// TIA Portal project "Mixing_Process" (V19)
// Mixing of two ingredients process

(* hardware
DEVICE "S7-1200 station_1"  S7-1200 Station
   slot 0: "Rack_0"  S7-1200 Rack  Rack  V1.0
   slot 1: "PLC_1"  CPU 1212C AC/DC/Rly  6ES7 212-1BE40-0XB0  V4.6
DEVICE "HMI_1"  TP1200 Comfort
   slot 0: "HMI_1"  TP1200 Comfort  6AV2 124-0MC01-0AX0  17.0.0.0
   slot 1: "HMI_RT_1"  TP1200 Comfort  6AV2 124-0MC01-0AX0  17.0.0.0
   slot 5: "HMI_1.IE_CP_1"  PROFINET Interface  17.0.0.0
      slot 1: "PROFINET Interface_1"  PROFINET Interface
         slot 1: "Port_1"  Port
         slot 2: "Port_2"  Port
   slot 7: "HMI_1.MPI/DP_CP_1"  MPI/DP Interface  17.0.0.0
*)

// ===== PLC "PLC_1"  CPU 1212C AC/DC/Rly =====

VAR_GLOBAL   // PLC tag table "Inputs"
   "E_Stop" AT %I0.0 : Bool;   // Stop mushroom
   "Pb_Stop" AT %I0.1 : Bool;   // Pushbutton Stop
   "Pb_Start" AT %I0.2 : Bool;   // Pushbutton Start
   "Tank_Empty_Level" AT %I0.3 : Bool;   // Empty level sensor, NO logic
   "Level_A" AT %I0.4 : Bool;   // Level for liquid A, NO logic
   "Level_B" AT %I0.5 : Bool;   // Level for liquid B, NO logic
   "Thermal_Fault" AT %I0.6 : Bool;   // Thermal fault from thermal relay
   "Temp_Alm" AT %I0.7 : Bool;   // Temperature alarm from control temperature
   "Tag_1" AT %M0.0 : Bool;
END_VAR

VAR_GLOBAL   // PLC tag table "Outputs"
   "Motor_Mixer" AT %Q0.0 : Bool;   // Motor mixer
   "Valve_A" AT %Q0.1 : Bool;   // Valve liquid A
   "Valve_B" AT %Q0.2 : Bool;   // Valve liquid B
   "Temp_Relay" AT %Q0.4 : Bool;   // Control relay for temperature signal
   "Valve_C" AT %Q0.5 : Bool;   // Discharge Valve
END_VAR

// folder: DB

DATA_BLOCK "DATA"   // DB1
TITLE = Data blocks for functions
{ S7_Optimized_Access := 'TRUE' }
AUTHOR : Stiven Perez Mora
VERSION : 0.1
   VAR
      Start_Stop : Bool;
      Q_TimeDischarge : Bool;
      E_Discharge : Int;
      Active_Valve_C : Bool;
      E_Active_Valve_C : Bool;
      E_Stop : Bool;
      Pb_Start : Bool;
   END_VAR
BEGIN
END_DATA_BLOCK

DATA_BLOCK "HMI_Data"   // DB4
{ S7_Optimized_Access := 'TRUE' }
VERSION : 0.1
   VAR
      Start_HMI : Bool;
      Stop_HMI : Bool;
      Valve_A : Bool;
      Level_A : Bool;
      Valve_B : Bool;
      Level_B : Bool;
      Valve_C : Bool;
      Motor_Mixer : Bool;
      Temp_Relay : Bool;
      PT_Mixing : Time;   // Miliseconds timer mix
      PT_M_Mxing : Time;   // Minutes timer mix
      ET_Mixing : Time;   // Miliseconds elapsed time
      ET_Mixing_S : Time;   // Seconds elapsed time
      Empty_Level : Bool;
      Empty_Field_Time : Bool;   // Ambar text alert, input mix time
   END_VAR
BEGIN
END_DATA_BLOCK

// folder: System blocks/Program resources

DATA_BLOCK "TimeToWamUp"   // DB2
{ S7_Optimized_Access := 'TRUE' }
AUTHOR : Simatic
FAMILY : IEC
NAME : IEC_TMR
VERSION : 1.0
// stored: InstanceOfName IEC_TIMER
"IEC_TIMER"
BEGIN
END_DATA_BLOCK

DATA_BLOCK "TimeToMixing"   // DB3
{ S7_Optimized_Access := 'TRUE' }
AUTHOR : Simatic
FAMILY : IEC
NAME : IEC_TMR
VERSION : 1.0
// stored: InstanceOfName IEC_TIMER
"IEC_TIMER"
BEGIN
END_DATA_BLOCK

DATA_BLOCK "MixingTime"   // DB5
{ S7_Optimized_Access := 'TRUE' }
AUTHOR : Simatic
FAMILY : IEC
NAME : IEC_TMR
VERSION : 1.0
// stored: InstanceOfName IEC_TIMER
"IEC_TIMER"
BEGIN
END_DATA_BLOCK

// folder: (top level)

ORGANIZATION_BLOCK "Main"   // OB1, LAD, ProgramCycle
TITLE = "Main Program Sweep (Cycle)"
{ S7_Optimized_Access := 'TRUE' }
VERSION : 0.1
   VAR_INPUT
      Initial_Call : Bool;   // Initial call of this OB
      Remanence : Bool;   // =True, if remanent data are available
   END_VAR
BEGIN

REGION Network 1: Block Start or Stop all process
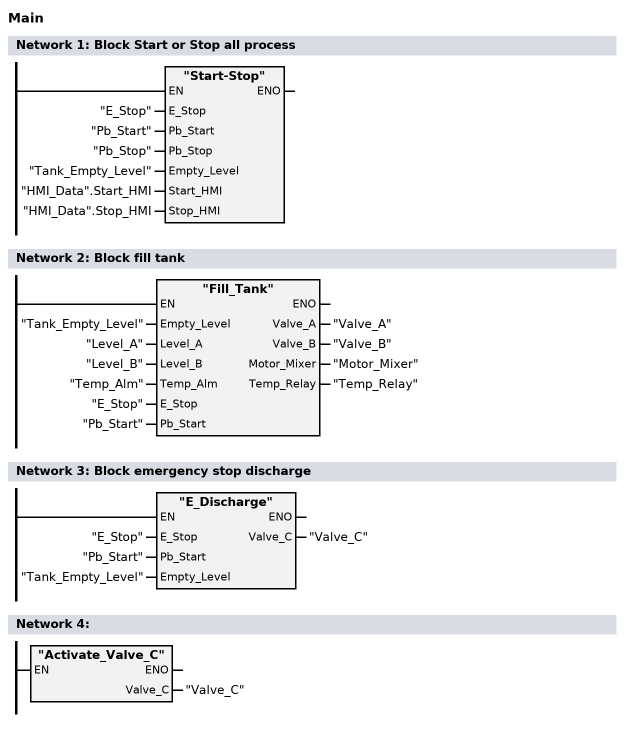
   RUNG wire#powerrail
      "Start-Stop"(E_Stop := "E_Stop", Pb_Start := "Pb_Start", Pb_Stop := "Pb_Stop", Empty_Level := "Tank_Empty_Level", Start_HMI := "HMI_Data".Start_HMI, Stop_HMI := "HMI_Data".Stop_HMI)
   END_RUNG
   // the same network as SCL:
   "Start-Stop"(E_Stop := "E_Stop",
                Pb_Start := "Pb_Start",
                Pb_Stop := "Pb_Stop",
                Empty_Level := "Tank_Empty_Level",
                Start_HMI := "HMI_Data".Start_HMI,
                Stop_HMI := "HMI_Data".Stop_HMI);
END_REGION

REGION Network 2: Block fill tank
   RUNG wire#powerrail
      "Fill_Tank"(Empty_Level := "Tank_Empty_Level", Level_A := "Level_A", Level_B := "Level_B", Temp_Alm := "Temp_Alm", E_Stop := "E_Stop", Pb_Start := "Pb_Start", Valve_A => "Valve_A", Valve_B => "Valve_B", Motor_Mixer => "Motor_Mixer", Temp_Relay => "Temp_Relay")
   END_RUNG
   // the same network as SCL:
   "Fill_Tank"(Empty_Level := "Tank_Empty_Level",
               Level_A := "Level_A",
               Level_B := "Level_B",
               Temp_Alm := "Temp_Alm",
               E_Stop := "E_Stop",
               Pb_Start := "Pb_Start",
               Valve_A => "Valve_A",
               Valve_B => "Valve_B",
               Motor_Mixer => "Motor_Mixer",
               Temp_Relay => "Temp_Relay");
END_REGION

REGION Network 3: Block emergency stop discharge
   RUNG wire#powerrail
      "E_Discharge"(E_Stop := "E_Stop", Pb_Start := "Pb_Start", Empty_Level := "Tank_Empty_Level", Valve_C => "Valve_C")
   END_RUNG
   // the same network as SCL:
   "E_Discharge"(E_Stop := "E_Stop",
                 Pb_Start := "Pb_Start",
                 Empty_Level := "Tank_Empty_Level",
                 Valve_C => "Valve_C");
END_REGION

REGION Network 4
   RUNG wire#powerrail
      "Activate_Valve_C"(Valve_C => "Valve_C")
   END_RUNG
   // the same network as SCL:
   "Activate_Valve_C"(Valve_C => "Valve_C");
END_REGION
END_ORGANIZATION_BLOCK

// folder: FC

FUNCTION "Start-Stop" : Void   // FC1, LAD
TITLE = Start stop process
{ S7_Optimized_Access := 'TRUE' }
AUTHOR : Stiven Perez Mora
VERSION : 0.1
// Conditions to active or deactive all process
   VAR_INPUT
      E_Stop : Bool;
      Pb_Start : Bool;
      Pb_Stop : Bool;
      Empty_Level : Bool;
      Start_HMI : Bool;
      Stop_HMI : Bool;
   END_VAR
BEGIN

REGION Network 1: Start Process
   // Conditions to start all process, initial conditions are, tank must be empty and operator must set the time for mixing, if mix time is equal to 0, the process will dont start
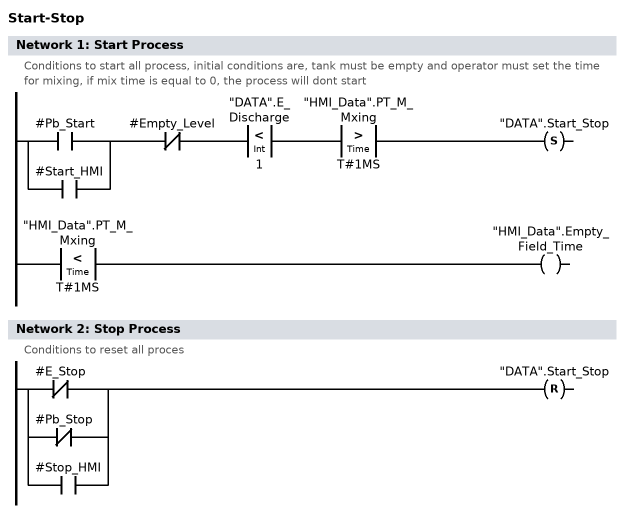
   RUNG wire#powerrail
      Contact( #Pb_Start )
      wire#w1
      I_Contact( #Empty_Level )
      { S7_Templates := "SrcType := Int" } LT_Contact(in1 := "DATA".E_Discharge, in2 := 1)
      { S7_Templates := "SrcType := Time" } GT_Contact(in1 := "HMI_Data".PT_M_Mxing, in2 := T#1MS)
      S_Coil( "DATA".Start_Stop )
   END_RUNG
   RUNG wire#powerrail
      Contact( #Start_HMI )
   END_RUNG wire#w1
   RUNG wire#powerrail
      { S7_Templates := "SrcType := Time" } LT_Contact(in1 := "HMI_Data".PT_M_Mxing, in2 := T#1MS)
      Coil( "HMI_Data".Empty_Field_Time )
   END_RUNG
   // the same network as SCL:
   IF (#Pb_Start OR #Start_HMI) AND NOT #Empty_Level AND ("DATA".E_Discharge < 1) AND ("HMI_Data".PT_M_Mxing > T#1MS) THEN
       "DATA".Start_Stop := TRUE;
   END_IF;
   "HMI_Data".Empty_Field_Time := "HMI_Data".PT_M_Mxing < T#1MS;
END_REGION

REGION Network 2: Stop Process
   // Conditions to reset all proces
   RUNG wire#powerrail
      I_Contact( #E_Stop )
      wire#w1
      R_Coil( "DATA".Start_Stop )
   END_RUNG
   RUNG wire#powerrail
      I_Contact( #Pb_Stop )
   END_RUNG wire#w1
   RUNG wire#powerrail
      Contact( #Stop_HMI )
   END_RUNG wire#w1
   // the same network as SCL:
   IF NOT #E_Stop OR NOT #Pb_Stop OR #Stop_HMI THEN "DATA".Start_Stop := FALSE; END_IF;
END_REGION
END_FUNCTION

FUNCTION "Fill_Tank" : Void   // FC2, LAD
TITLE = Fill Tank for mixing process
{ S7_Optimized_Access := 'TRUE' }
AUTHOR : Stiven Perez Mora
VERSION : 0.1
   VAR_INPUT
      Empty_Level : Bool;
      Level_A : Bool;
      Level_B : Bool;
      Temp_Alm : Bool;
      E_Stop : Bool;
      Pb_Start : Bool;
   END_VAR
   VAR_OUTPUT
      Valve_A : Bool;
      Valve_B : Bool;
      Motor_Mixer : Bool;
      Temp_Relay : Bool;
   END_VAR
BEGIN

REGION Network 1: Convert time from mixing timer
   // Convert elapsed time millisenconds to seconds and preset time
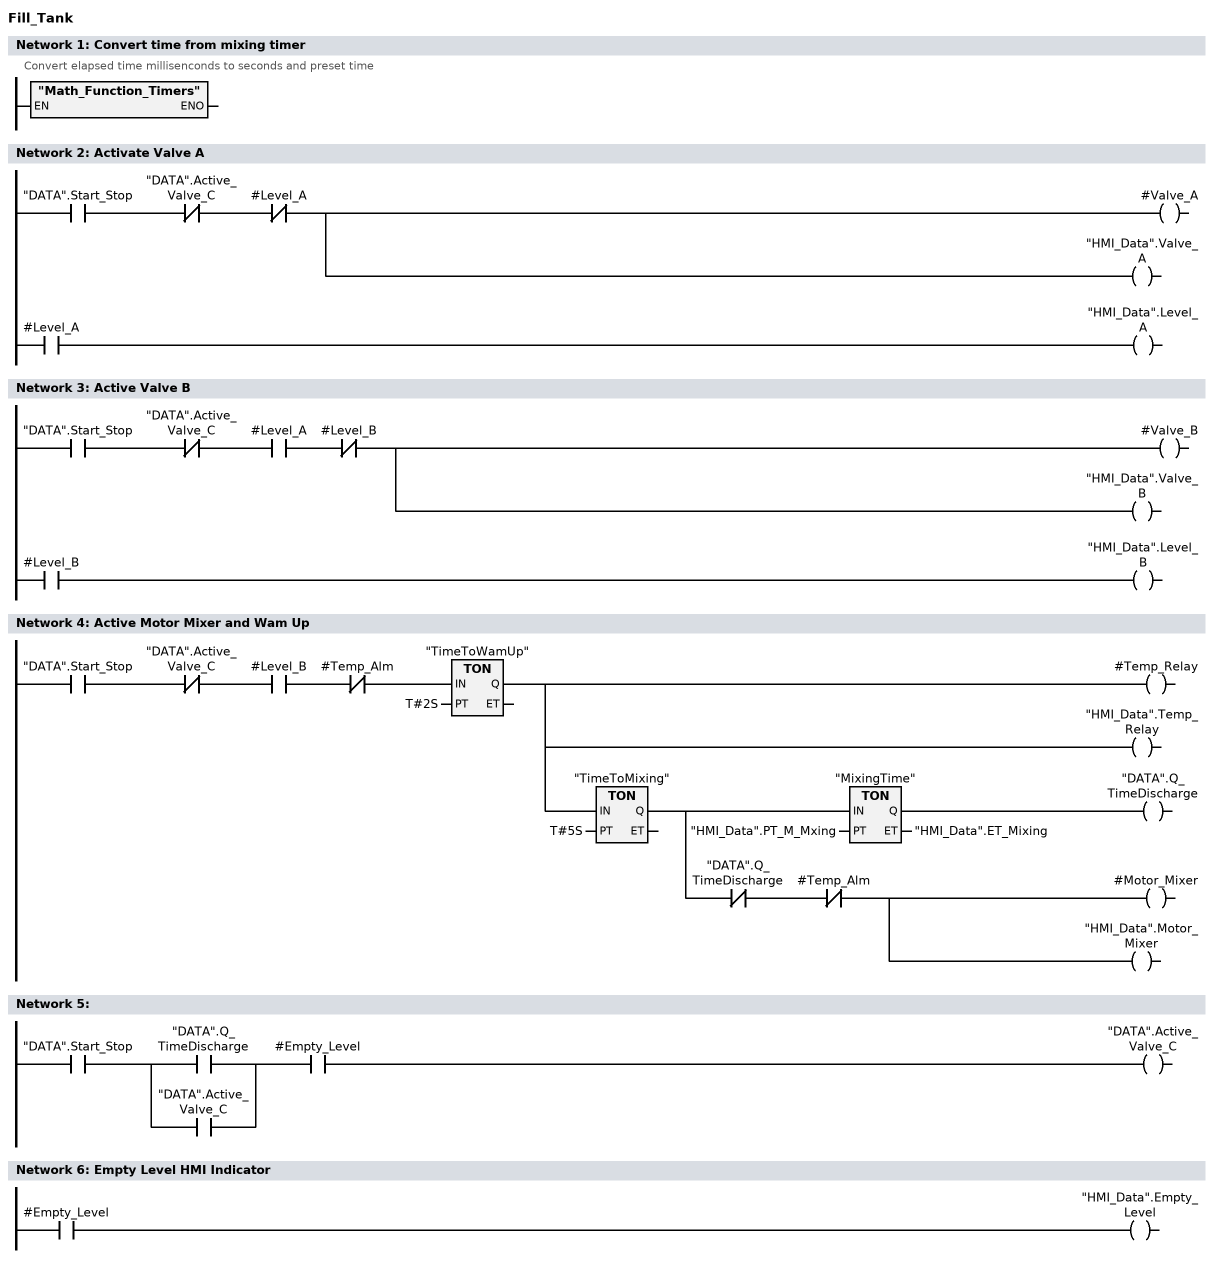
   RUNG wire#powerrail
      "Math_Function_Timers"()
   END_RUNG
   // the same network as SCL:
   "Math_Function_Timers"();
END_REGION

REGION Network 2: Activate Valve A
   RUNG wire#powerrail
      Contact( "DATA".Start_Stop )
      I_Contact( "DATA".Active_Valve_C )
      I_Contact( #Level_A )
      wire#w1
      Coil( #Valve_A )
   END_RUNG
   RUNG wire#w1
      Coil( "HMI_Data".Valve_A )
   END_RUNG
   RUNG wire#powerrail
      Contact( #Level_A )
      Coil( "HMI_Data".Level_A )
   END_RUNG
   // the same network as SCL:
   #Valve_A := "DATA".Start_Stop AND NOT "DATA".Active_Valve_C AND NOT #Level_A;
   "HMI_Data".Valve_A := #Valve_A;
   "HMI_Data".Level_A := #Level_A;
END_REGION

REGION Network 3: Active Valve B
   RUNG wire#powerrail
      Contact( "DATA".Start_Stop )
      I_Contact( "DATA".Active_Valve_C )
      Contact( #Level_A )
      I_Contact( #Level_B )
      wire#w1
      Coil( #Valve_B )
   END_RUNG
   RUNG wire#w1
      Coil( "HMI_Data".Valve_B )
   END_RUNG
   RUNG wire#powerrail
      Contact( #Level_B )
      Coil( "HMI_Data".Level_B )
   END_RUNG
   // the same network as SCL:
   #Valve_B := "DATA".Start_Stop AND NOT "DATA".Active_Valve_C AND #Level_A AND NOT #Level_B;
   "HMI_Data".Valve_B := #Valve_B;
   "HMI_Data".Level_B := #Level_B;
END_REGION

REGION Network 4: Active Motor Mixer and Wam Up
   "TimeToWamUp".TON(IN := "DATA".Start_Stop AND NOT "DATA".Active_Valve_C AND #Level_B AND NOT #Temp_Alm,
                     PT := T#2S);
   #Temp_Relay := "TimeToWamUp".Q;
   "HMI_Data".Temp_Relay := "TimeToWamUp".Q;
   "TimeToMixing".TON(IN := "TimeToWamUp".Q, PT := T#5S);
   "MixingTime".TON(IN := "TimeToMixing".Q, PT := "HMI_Data".PT_M_Mxing, ET => "HMI_Data".ET_Mixing);
   "DATA".Q_TimeDischarge := "MixingTime".Q;
   #Motor_Mixer := "TimeToMixing".Q AND NOT "DATA".Q_TimeDischarge AND NOT #Temp_Alm;
   "HMI_Data".Motor_Mixer := #Motor_Mixer;
END_REGION

REGION Network 5
   RUNG wire#powerrail
      Contact( "DATA".Start_Stop )
      wire#w1
      Contact( "DATA".Q_TimeDischarge )
      wire#w2
      Contact( #Empty_Level )
      Coil( "DATA".Active_Valve_C )
   END_RUNG
   RUNG wire#w1
      Contact( "DATA".Active_Valve_C )
   END_RUNG wire#w2
   // the same network as SCL:
   "DATA".Active_Valve_C := "DATA".Start_Stop AND ("DATA".Q_TimeDischarge OR "DATA".Active_Valve_C) AND #Empty_Level;
END_REGION

REGION Network 6: Empty Level HMI Indicator
   RUNG wire#powerrail
      Contact( #Empty_Level )
      Coil( "HMI_Data".Empty_Level )
   END_RUNG
   // the same network as SCL:
   "HMI_Data".Empty_Level := #Empty_Level;
END_REGION
END_FUNCTION

FUNCTION "Math_Function_Timers" : Void   // FC3, LAD
TITLE = Convert time from mixing timer
{ S7_Optimized_Access := 'TRUE' }
VERSION : 0.1
BEGIN

REGION Network 1: Input miliseconds time from HMI convert to Minutes
   // input field from HMI is equal to milliseconds, in this network millisencond are convert to minutes, the formula for convert milliseconds to minutes is multiply the data type from HMI field per 60.000
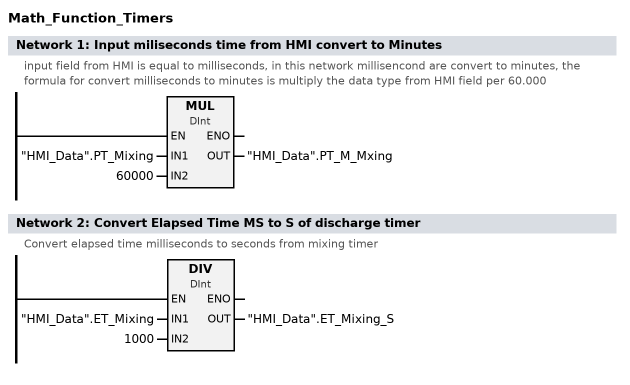
   RUNG wire#powerrail
      { S7_Templates := "SrcType := DInt" } Mul(in1 := "HMI_Data".PT_Mixing, in2 := 60000, out => "HMI_Data".PT_M_Mxing)
   END_RUNG
   // the same network as SCL:
   "HMI_Data".PT_M_Mxing := "HMI_Data".PT_Mixing * 60000;
END_REGION

REGION Network 2: Convert Elapsed Time MS to S of discharge timer
   // Convert elapsed time milliseconds to seconds from mixing timer
   RUNG wire#powerrail
      { S7_Templates := "SrcType := DInt" } Div(in1 := "HMI_Data".ET_Mixing, in2 := 1000, out => "HMI_Data".ET_Mixing_S)
   END_RUNG
   // the same network as SCL:
   "HMI_Data".ET_Mixing_S := "HMI_Data".ET_Mixing / 1000;
END_REGION
END_FUNCTION

FUNCTION "E_Discharge" : Void   // FC4, LAD
{ S7_Optimized_Access := 'TRUE' }
VERSION : 0.1
   VAR_INPUT
      E_Stop : Bool;
      Pb_Start : Bool;
      Empty_Level : Bool;
   END_VAR
   VAR_OUTPUT
      Valve_C : Bool;
   END_VAR
   VAR_TEMP   // added for the SCL form of the ladder/FBD networks
      _w1 : Bool;
      _w2 : Bool;
   END_VAR
BEGIN

REGION Network 1: Counter emergency stop pushed
   // if emergency stop has been pushed, the counter variable discharge increase 1, if counter variable is equal to 1 the valve C will activate but the tank must be filled, when the level decrease, the empty level sensor deactivate valve C and enable push button start for restart counter variable and start process
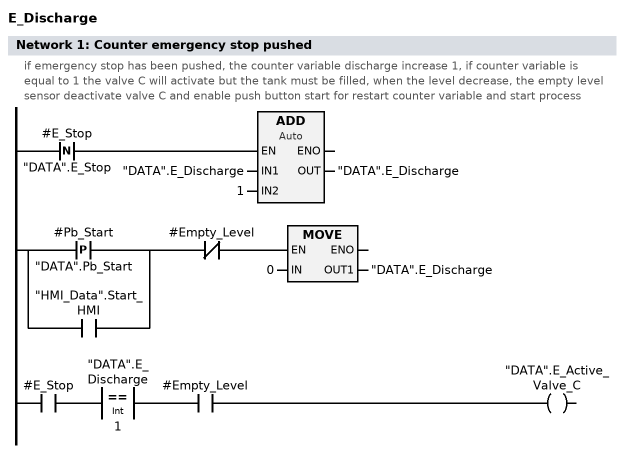
   RUNG wire#powerrail
      N_Contact(operand := #E_Stop, bit := "DATA".E_Stop)
      Add(in1 := "DATA".E_Discharge, in2 := 1, out => "DATA".E_Discharge)
   END_RUNG
   RUNG wire#powerrail
      P_Contact(operand := #Pb_Start, bit := "DATA".Pb_Start)
      wire#w1
      I_Contact( #Empty_Level )
      Move(in := 0, out1 => "DATA".E_Discharge)
   END_RUNG
   RUNG wire#powerrail
      Contact( "HMI_Data".Start_HMI )
   END_RUNG wire#w1
   RUNG wire#powerrail
      Contact( #E_Stop )
      { S7_Templates := "SrcType := Int" } EQ_Contact(in1 := "DATA".E_Discharge, in2 := 1)
      Contact( #Empty_Level )
      Coil( "DATA".E_Active_Valve_C )
   END_RUNG
   // the same network as SCL:
   #_w1 := NOT #E_Stop AND "DATA".E_Stop;   // falling edge of #E_Stop
   "DATA".E_Stop := #E_Stop;
   IF #_w1 THEN "DATA".E_Discharge := "DATA".E_Discharge + 1; END_IF;
   #_w2 := #Pb_Start AND NOT "DATA".Pb_Start;   // rising edge of #Pb_Start
   "DATA".Pb_Start := #Pb_Start;
   IF (#_w2 OR "HMI_Data".Start_HMI) AND NOT #Empty_Level THEN "DATA".E_Discharge := 0; END_IF;
   "DATA".E_Active_Valve_C := #E_Stop AND ("DATA".E_Discharge = 1) AND #Empty_Level;
END_REGION
END_FUNCTION

FUNCTION "Activate_Valve_C" : Void   // FC5, LAD
{ S7_Optimized_Access := 'TRUE' }
VERSION : 0.1
   VAR_OUTPUT
      Valve_C : Bool;
   END_VAR
BEGIN

REGION Network 1: Discharge Valve
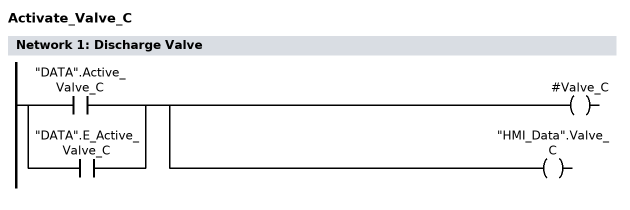
   RUNG wire#powerrail
      Contact( "DATA".Active_Valve_C )
      wire#w1
      Coil( #Valve_C )
   END_RUNG
   RUNG wire#powerrail
      Contact( "DATA".E_Active_Valve_C )
   END_RUNG wire#w1
   RUNG wire#w1
      Coil( "HMI_Data".Valve_C )
   END_RUNG
   // the same network as SCL:
   #Valve_C := "DATA".Active_Valve_C OR "DATA".E_Active_Valve_C;
   "HMI_Data".Valve_C := #Valve_C;
END_REGION
END_FUNCTION

// ===== library types =====

// folder: LGF/1 Date and timer operations

FUNCTION "LGF_GetCalendarDay" : DInt   // FC10028, SCL
TITLE = LGF_GetCalendarDay
{ S7_Optimized_Access := 'TRUE' }
AUTHOR : Siemens_Digital_Industry
FAMILY : LGF
NAME : LGF_GetCalendarDay
// This function uses the specified date to calculate the number of days that have passed since the beginning of the year (1st January).
// 
// The function is used in the functions “LGF_GetCalendarWeek_ISO” and “LGF_GetCalendarWeek_US”.
// Diese Funktion berechnet aus dem vorgegebenen Datum die Anzahl der Tage, die seit dem Anfang des Jahres vergangen sind (1. Januar).
// 
// Die Funktion wird in den Funktionen "LGF_GetCalendarWeek_ISO" und "LGF_GetCalendarWeek_US" verwendet.
   VAR_INPUT
      "date" : DTL;   // Date for the calculation of the calendar days since 1 January. / Datum für die Berechnung der vergangenen Kalendertagen seit dem 01. Januar
   END_VAR
   VAR_OUTPUT
      error : Bool;   // FALSE: No error / TRUE: An error occurred during the execution of the FB / FALSE: Kein Fehler / TRUE: Während der Ausführung des FB ist ein Fehler aufgetreten
      status : Word;   // 16#0000-16#7FFF: Status of the FB / 16#8000-16#FFFF: Error identification (see following Table) / 16#0000-16#7FFF: Status des FB / 16#8000-16#FFFF: Fehleridentifikation (siehe folgende Tabelle)
   END_VAR
   VAR_TEMP
      tempDaysPassed : DInt;   // Temp tag for the number of days past / Temp Variable für die Anzahl der vergangenen Tage
      tempDate : DTL;   // Temp variable to store date for calculations / Temp Variable um Datum für Berechung zwischen zu speichern
   END_VAR
   // Ret_Val : Days past since January 1st. / Vergangene Tage seit 1. Januar.
   VAR CONSTANT
      FIRST_DAY : USInt := 1;   // 1st of a month / 1. Tag eines Monats
      LAST_DAY : USInt := 31;   // 31st of a month / 31. Tag eines Monats
      JANUARY : USInt := 1;   // Month number for January / Monatsnumer Januar
      DECEMBER : USInt := 12;   // Month number for December / Monatsnummer Dezember
      TIME_ZERO_FORCE_UPDATE : Time := t#0d;   // By adding zero an update of DTL Tag is forced and auto checks are applied / Durch die Addition von "0" wird ein Update üder den Zeitstemple erstellt und ebenfalls auf gültigkeit geprüft.
      ONE_DAY : DInt := 1;   // One single day for incrementing / Ein Tag für inkrementierungen
      STATUS_NO_ERROR : Word := 16#0000;   // Status: no error occurred / Status: kein Fehler aufgetreten
      ERR_LIM_DATE : Word := 16#8201;   // Date out of the range, has to be greater than <1970-01-01 ; 2262-04-11> / Datum ausserhalb des gültigen Bereiches, es muss nach dem <1970-01-01 ; 2262-04-11> liegen
   END_VAR
BEGIN
   REGION BLOCK INFO HEADER
     //===============================================================================
     // SIEMENS AG / (c)Copyright 2019
     //-------------------------------------------------------------------------------
     // Title:            LGF_GetCalendarDay
     // Comment/Function: This function calculates for a date the passed days since 1st January.
     // Library/Family:   LGF(Library General Functions)
     // Author:           Siemens Digital Industry Support
     // Tested with:      S7-PLCSIM Advanced V2.0 SP1
     // Engineering:      TIA Portal V15.1
     // Restrictions:     ENO disabled - error handling done with error and status
     // Requirements:     PLC (S7-1200 / S7-1500)
     //-------------------------------------------------------------------------------
     // Change log table:
     // Version  | Date       | Expert in charge       | Changes applied
     //----------|------------|------------------------|------------------------------
     // 01.00.00 16.07.2019  Simatic Systems Support
     //                      First release
     //                      ENO used for internal error handling, interface has error and status
     //                      temp tag naming, insert constant
     // 03.00.00 23.04.2020  Simatic Systems Support
     //                      Set version to V3.0.0, harmonize the version of the whole library
     // 03.00.01 19.01.2020  Simatic Systems Support
     //                      Insert documentation
     //=============================================================================
   END_REGION BLOCK INFO HEADER

   REGION INITIALISATION
     #tempDate := #date;
     #tempDaysPassed := 0;
   END_REGION

   REGION COUNT DAYS
     // Check #date
     // adding zero forces the PLC to update the tag and eno check
     #tempDate := #tempDate + #TIME_ZERO_FORCE_UPDATE;
     IF ENO = FALSE THEN
       #error := TRUE;
       #status := #ERR_LIM_DATE;
       #LGF_GetCalendarDay := #tempDaysPassed;
       RETURN;
     END_IF;

     // Weekday of 1st January in the current year
     #tempDate.MONTH := #JANUARY;
     #tempDate.DAY := #FIRST_DAY;
     // adding zero forces the PLC to update the tag
     // in this case especially the weekday
     #tempDate := #tempDate + #TIME_ZERO_FORCE_UPDATE;

     // Days passed in the year since 1st January, "date" included
     #tempDaysPassed := DATE_TO_DINT(DTL_TO_DATE(#date)) - DATE_TO_DINT(DTL_TO_DATE(#tempDate)) + #ONE_DAY;
   END_REGION

   REGION OUTPUTS
     #error := FALSE;
     #status := #STATUS_NO_ERROR;
     #LGF_GetCalendarDay := #tempDaysPassed;

     // ENO is not used, forced to TRUE
     ENO := TRUE;
   END_REGION
END_FUNCTION

(* ===== HMI "HMI_RT_1" =====
system functions are stored by id; their names below are inferred from use
connection "HMI_Connection_3": ETHERNET, S7_1200_OMS

HMI tags "DATA"
   "Start" : Bool = PLC HMI_Data.Start_HMI AT %I0.2, 100 ms
   "Stop" : Bool = PLC HMI_Data.Stop_HMI AT %I0.1, 100 ms
   "Valve_A" : Bool = PLC HMI_Data.Valve_A AT %DB1.DBX0.0, 100 ms
   "Valve_B" : Bool = PLC HMI_Data.Valve_B AT %DB1.DBX0.0, 100 ms
   "Valve_C" : Bool = PLC HMI_Data.Valve_C AT %DB1.DBX0.0, 100 ms
   "Motor_Mixer" : Bool = PLC HMI_Data.Motor_Mixer AT %DB1.DBX0.0, 100 ms
   "Temp_Relay" : Bool = PLC HMI_Data.Temp_Relay AT %DB1.DBX0.0, 100 ms
   "ET_Mixing" : Time = PLC HMI_Data.ET_Mixing_S, 100 ms
   "Level_A" : Bool = PLC HMI_Data.Level_A AT %I0.4, 100 ms
   "Level_B" : Bool = PLC HMI_Data.Level_B AT %I0.5, 100 ms
   "Empty_Tank" : Bool = PLC HMI_Data.Empty_Level AT %I0.3, 100 ms
   "PT_Mixing" : Time = PLC HMI_Data.PT_Mixing AT %DB1.DBX0.0, 100 ms
   "Empty_Field_Time" : Bool = PLC HMI_Data.Empty_Field_Time AT %DB1.DBW0, 1 s
   "Start_Stop" : Bool = PLC DATA.Start_Stop AT %DB1.DBX0.0, 1 s

Template "Template_1" 1280x740
   Button "Exit" at 1200,679 size 78x59; TextOff 'Exit'; PictureOff "ExitRuntime_TP1200_Comfort_TR"; PictureOn "ExitRuntime_TP1200_Comfort_TR"
      on Release: StopRuntime(0)
   Button "Template_Button" at 1120,679 size 78x59; TextOff 'Text'
   Button "Template_Button_1" at 1040,679 size 78x59; TextOff 'Text'
   Button "Template_Button_2" at 960,679 size 78x59; TextOff 'Text'
   Button "Template_Button_3" at 880,679 size 78x59; TextOff 'Text'
   Button "Template_Button_4" at 800,679 size 78x59; TextOff 'Text'
   Button "Template_Button_5" at 720,679 size 78x59; TextOff 'Text'
   Button "Template_Button_6" at 640,679 size 78x59; TextOff 'Text'
   Button "Template_Button_7" at 561,679 size 78x59; TextOff 'Text'
   Button "Template_Button_8" at 481,679 size 78x59; TextOff 'Text'
   Button "Template_Button_9" at 401,679 size 78x59; TextOff 'Text'
   Button "Template_Button_10" at 321,679 size 78x59; TextOff 'Text'
   Button "Template_Button_11" at 241,679 size 78x59; TextOff 'Text'
   Button "Template_Button_12" at 161,679 size 78x59; TextOff 'Text'
   Button "Template_Button_13" at 81,679 size 78x59; TextOff 'Text'
   Button "Start screen" at 1,679 size 78x59; TextOff 'Start screen'; PictureOff "NavigateHome_TP1200_Comfort_TR"; PictureOn "NavigateHome_TP1200_Comfort_TR"
      on Release: ActivateScreen("Root screen", 0)
   AlarmView "Alarm view_Unacknowledged" at 0,0 size 1280x23

screen "Root screen" 1280x740, template "Template_1"
   GraphicView "Graphic view_1" at 457,173 size 370x354; Picture "Graphic_1"
   GraphicView "Graphic view_3" at 628,545 size 37x33; Picture "Graphic_6"
   GraphicView "Graphic view_6" at 654,554 size 235x28; Picture "Graphic_7"
   GraphicView "Graphic view_7" at 621,521 size 31x28; Picture "Graphic_5"
   GraphicView "Graphic view_8" at 262,150 size 125x28; Picture "Graphic_7"
   GraphicView "Graphic view_9" at 879,149 size 125x28; Picture "Graphic_7"
   GraphicView "Graphic view_10" at 763,149 size 59x28; Picture "Graphic_7"
   GraphicView "Graphic view_11" at 445,149 size 59x28; Picture "Graphic_7"
   GraphicView "Graphic view_12" at 500,155 size 43x33; Picture "Graphic_9"
   GraphicView "Graphic view_13" at 730,155 size 37x33; Picture "Graphic_10"
   GraphicView "Graphic view_14" at 585,67 size 107x284; Picture "Graphic_11"
      Visibility <- "Motor_Mixer"
   GraphicView "Graphic view_15" at 557,323 size 163x139; Picture "Graphic_15"
      Visibility <- "Temp_Relay"
   TextField "Text field_1" at 835,111 size 30x25; Text 'VB'
      Appearance <- "Valve_B"
   TextField "Text field_2" at 402,110 size 30x25; Text 'VA'
      Appearance <- "Valve_A"
   TextField "Text field_3" at 896,515 size 29x25; Text 'VC'
      Appearance <- "Valve_C"
   GraphicView "Graphic view_16" at 942,554 size 59x28; Picture "Graphic_7"
   Button "Button_1" at 57,222 size 171x64; TextOff 'START'
      on Press: function_b14e0dd5("Start", 0)
      Appearance <- "Start_Stop"
      ProcessValue <- "Start_Stop"
   Button "Button_2" at 56,326 size 171x64; TextOff 'STOP'
      on Press: function_b14e0dd5("Stop", 0)
      Appearance <- "Stop"
   GraphicView "Graphic view_2" at 586,68 size 105x283; Picture "Graphic_21"
      Visibility <- "Motor_Mixer"
   IOField "I/O field_1" at 70,541 size 93x40; FormatPattern 99
      ProcessValue <- "PT_Mixing"
   Rectangle "Rectangle_1" at 1039,243 size 155x62
      Visibility <- "Level_A"
   TextField "Text field_4" at 1066,256 size 102x34; Text 'Level A'
      Visibility <- "Level_A"
   Rectangle "Rectangle_2" at 1039,328 size 155x62
      Visibility <- "Level_B"
   TextField "Text field_5" at 1066,341 size 102x34; Text 'Level B'
      Visibility <- "Level_B"
   Rectangle "Rectangle_3" at 1039,416 size 155x62
      Visibility <- "Empty_Tank"
   TextField "Text field_6" at 1046,430 size 152x32; Text 'Tank Empty'
      Visibility <- "Empty_Tank"
   TextField "Text field_7" at 51,501 size 163x27; Text 'Enter Mix Time'
      Appearance <- "Empty_Field_Time"
   IOField "I/O field_2" at 301,541 size 101x39; FormatPattern 9999
      ProcessValue <- "ET_Mixing"
   TextField "Text field_8" at 290,500 size 133x27; Text 'Mixing Time'
   GraphicView "Graphic view_19" at 879,543 size 67x43; Picture "Graphic_25"
      Visibility <- "Valve_C"
   GraphicView "Graphic view_18" at 818,138 size 67x43; Picture "Graphic_25"
      Visibility <- "Valve_B"
   GraphicView "Graphic view_20" at 382,138 size 67x43; Picture "Graphic_25"
      Visibility <- "Valve_A"
   GraphicView "Graphic view_21" at 878,542 size 69x46; Picture "Graphic_26"
      Visibility <- "Valve_C"
   GraphicView "Graphic view_22" at 381,137 size 69x46; Picture "Graphic_26"
      Visibility <- "Valve_A"
   GraphicView "Graphic view_23" at 817,137 size 69x46; Picture "Graphic_26"
      Visibility <- "Valve_B"
   TextField "Text field_9" at 169,550 size 39x25; Text 'Min'
   TextField "Text field_10" at 110,241 size 65x25; Text 'START'
      Visibility <- "Start_Stop"
   TextField "Text field_11" at 1050,210 size 136x25; Text 'Level Sensors'
   TextField "Text field_12" at 407,549 size 38x25; Text 'Sec'
   GraphicView "Graphic view_25" at 741,559 size 23x20; Picture "right-arrow"
      Appearance <- "Valve_C"
      Visibility <- "Valve_C"
   GraphicView "Graphic view_26" at 960,559 size 23x20; Picture "right-arrow"
      Appearance <- "Valve_C"
      Visibility <- "Valve_C"
   GraphicView "Graphic view_27" at 635,559 size 23x20; Picture "right-arrow"
      Appearance <- "Valve_C"
      Visibility <- "Valve_C"
   GraphicView "Graphic view_4" at 312,155 size 23x20; Picture "right-arrow"
      Visibility <- "Valve_A"
      Appearance <- "Valve_A"
   GraphicView "Graphic view_24" at 487,154 size 23x20; Picture "right-arrow"
      Visibility <- "Valve_A"
      Appearance <- "Valve_A"
   GraphicView "Graphic view_5" at 759,152 size 29x22; Picture "left-arrow"
      Visibility <- "Valve_B"
      Appearance <- "Valve_B"
   GraphicView "Graphic view_17" at 919,152 size 29x22; Picture "left-arrow"
      Visibility <- "Valve_B"
      Appearance <- "Valve_B"
   GraphicView "Graphic view_28" at 835,559 size 23x20; Picture "right-arrow"
      Appearance <- "Valve_C"
      Visibility <- "Valve_C"
*)